(* Logix 5000 project; controller FV vendor 1 type 14 code 217 rev 31.11; software revision 31.00 *)

TASK _1Sec (periodic, rate 1000 ms, priority 10, watchdog 500 ms) : _1Second
TASK MainTask (continuous, watchdog 500 ms) : First_Task, FV_Common, FR_Common, Last_Task

MODULES
   Local : vendor 1 type 14 code 217 (5069 0, rev 31.11)
      MV : vendor 1 type 14 code 217 (Ethernet 192.168.20.32, rev 31.1)
      Remote_IO : vendor 1 type 12 code 298 (Ethernet 192.168.1.1, rev 1.1)
          : vendor 1 type 7 code 82 (Compact 6, rev 1.1, Input RPI 20 ms)
          : vendor 1 type 7 code 76 (Compact 7, rev 1.1, Input RPI 20 ms)
          : vendor 1 type 10 code 47 (Compact 8, rev 1.1, Output RPI 80 ms)
          : 1769-OW16 (Compact 1, rev 1.1, Output RPI 20 ms)
          : 1769-OW16 (Compact 3, rev 1.1, Output RPI 20 ms)
          : 1769-IF8 (Compact 13, rev 1.1, Output RPI 80 ms)
          : 1769-OW16 (Compact 4, rev 1.1, Output RPI 20 ms)
          : 1769-IF8 (Compact 11, rev 1.1, Output RPI 80 ms)
          : 1769-IF8 (Compact 10, rev 1.1, Output RPI 80 ms)
          : 1769-OW16 (Compact 2, rev 1.1, Output RPI 20 ms)
          : 1769-OW16 (Compact 5, rev 1.1, Output RPI 20 ms)
          : 1769-IF8 (Compact 12, rev 1.1, Output RPI 80 ms)
          : vendor 1 type 7 code 79 (Compact 9, rev 3.1, Output RPI 20 ms)
      RIO_Rack_2 : vendor 1 type 12 code 298 (Ethernet 192.168.1.2, rev 1.1)
          : vendor 1 type 7 code 76 (Compact 6, rev 1.1, Input RPI 20 ms)
          : vendor 1 type 7 code 76 (Compact 3, rev 1.1, Input RPI 20 ms)
          : vendor 1 type 7 code 76 (Compact 4, rev 1.1, Input RPI 20 ms)
          : vendor 1 type 7 code 76 (Compact 7, rev 1.1, Input RPI 20 ms)
          : vendor 1 type 7 code 76 (Compact 9, rev 1.1, Input RPI 20 ms)
          : vendor 1 type 7 code 76 (Compact 10, rev 1.1, Input RPI 20 ms)
          : vendor 1 type 7 code 76 (Compact 12, rev 1.1, Input RPI 20 ms)
          : vendor 1 type 7 code 79 (Compact 8, rev 3.1, Output RPI 20 ms)
          : vendor 1 type 10 code 48 (Compact 1, rev 1.1, Output RPI 80 ms)
          : vendor 1 type 10 code 47 (Compact 2, rev 1.1, Output RPI 80 ms)
          : vendor 1 type 7 code 79 (Compact 5, rev 3.1, Output RPI 20 ms)
          : vendor 1 type 7 code 79 (Compact 11, rev 3.1, Output RPI 20 ms)
      RIO_Rack_3 : vendor 1 type 12 code 298 (Ethernet 192.168.1.3, rev 1.1)
          : 1769-IQ16 (Compact 1, rev 1.1, Input RPI 20 ms)
          : 1769-IQ16 (Compact 2, rev 1.1, Input RPI 20 ms)
          : 1769-OW16 (Compact 3, rev 1.1, Output RPI 20 ms)
END_MODULES

TYPE CHECKWORD_FLAGS :   // Checkword Flags
STRUCT
   AUTODRV : DINT;   // Auto-Drive Bit No.
   CLOSEDFB : DINT;   // Closed Feedback Bit No.
   OPENFB : DINT;   // Open Feedback Bit No.
   OUTPUT : DINT;   // Output Bit No.
   MANDRV : DINT;   // Manual Drive Bit No.
   MANUAL : DINT;   // Manual Control Bit No.
   CHECKOFF : DINT;   // Checking Off Bit No.
   TRIPPED : DINT;   // Tripped Bit No.
   FAULT : DINT;   // Fault Bit No.
   SIMFAIL : DINT;   // Simulate Failure Bit
   PREVSCAN : DINT;   // Previous Scan State
   FAULTLOGGED : DINT;   // Fault Logged Flag From Scada
   HIGHLIGHT : DINT;   // Highlight on Graphics
   RUNFB : DINT;   // Pump/Drive Run Feedback
   HEALTHYFB : DINT;   // Pump Healthy Feedback
   NOTTRIPPEDFB : DINT;   // Pump Not Tripped Feedback
   HEALTHYFAULTLOGGED : DINT;   // Pump Not Healthy Fault Logged
   TRIPPEDFAULTLOGGED : DINT;   // Pump Tripped Fault Logged
   INPUTSTATUS : DINT;   // Bit Number for Digital Input Status
   INPUTSTATUSDEBOUNCED : DINT;   // Bit Number For Debounced Input Status
   ANALOGSIMULATION : DINT;   // Bit Number For Analog Simulation Enabled, Used By FactoryTalk
END_STRUCT
END_TYPE

TYPE DateTime :
STRUCT
   Year : DINT;
   Month : DINT;
   Day : DINT;
   Hour : DINT;
   Minute : DINT;
   Second : DINT;
   Microsecond : DINT;
END_STRUCT
END_TYPE

TYPE PlantItem :   // Plant Item
STRUCT
   CW : DINT;   // Checkword
   CheckTime : DINT;   // Check Time
   CheckTimer : DINT;   // Check Time Timer
   DebounceTime : DINT;   // Debounce Time
   DebounceTimer : DINT;   // Debounce Timer
   DriveBits : DINT;   // Item Automatic Drive Bits
   Scaled : REAL;   // Analogue Value Scaled For Input/Output
   RawInput : REAL;   // Raw Input Copied for display On Factory Talk
END_STRUCT
END_TYPE

TYPE Process :   // Data Type For Processes
STRUCT
   Status : DINT;   // Process Current Status
   Step : DINT;   // Process Current Step
   Step_Timer : DINT;   // Current Step Timer
   Fault : DINT;   // Process Current Fault
   Cmd : DINT;   // Command From Scada
   Cmd_avail : DINT;   // Commands Available To Scada
   Cmd_ok : BOOL;   // Startup Command Is Valid Flag
   Cmd_reset : TIMER;   // Startup timer for Invalid Command
   Data_scada : REAL[50];   // Data from Scada
   Data_work : REAL[50];   // Working Data in use by PLC
   Drivebit : DINT;   // Bit Number to Drive Plant Items With
   MessageID : DINT;   // ID to pass with Events/Alarms to Scada
   Past_Prestart : BOOL;   // Flag Set to Indicate past pre start checks.
   Restart_Step : DINT;   // Step to go back to after Continue
END_STRUCT
END_TYPE

TYPE Route :
STRUCT
   CW : DINT;   // Checking Group CW
   CW_Itm : DINT;   // Checking Group Which Has Failed
   Operation : DINT;   // Checking Group Operation Reservation
END_STRUCT
END_TYPE

ADD_ON_INSTRUCTION DayOfWeek   (* revision 1.0 *)
VAR_INPUT
   Year : DINT; {required}
   Month : DINT; {required}
   Day : DINT; {required}
END_VAR
VAR_OUTPUT
   DOW_Output : DINT; {access Read Only, required}
END_VAR
VAR
   DOW_Day : DINT;
   DOW_Year : DINT;
   DOW_Temp00 : REAL;
   DOW_Century : DINT;
   DOW_Month : DINT;
   DOW_Temp01 : REAL;
   DOW_Temp02 : REAL;
   DOW_Temp03 : DINT;
   DOW_Temp04 : DINT;
   DOW_Temp05 : REAL;
   DOW_Temp06 : DINT;
   DOW_Temp07 : REAL;
   DOW_Temp08 : DINT;
   DOW_Temp09 : REAL;
   DOW_Temp10 : REAL;
   DOW_Temp11 : REAL;
   DOW_Temp12 : REAL;
   DOW_Temp13 : REAL;
   DOW_Temp14 : REAL;
   DOW_Temp15 : REAL;
END_VAR

ROUTINE Logic   (* ladder *)
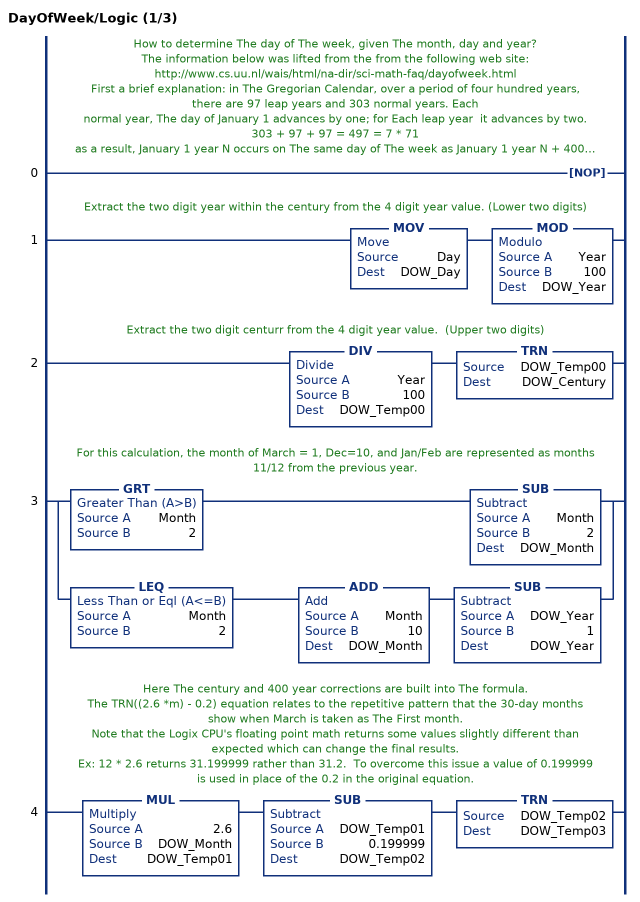
   // How to determine The day of The week, given The month, day and year?
   // The information below was lifted from the from the following web site: http://www.cs.uu.nl/wais/html/na-dir/sci-math-faq/dayofweek.html
   //    First a brief explanation: in The Gregorian Calendar, over a period of four hundred years, there are 97 leap years and 303 normal years. Each
   //  normal year, The day of January 1 advances by one; for Each leap year  it advances by two.
   //    303 + 97 + 97 = 497 = 7 * 71
   //    as a result, January 1 year N occurs on The same day of The week as January 1 year N + 400. Because The leap year pattern also recurs with a four hundred year cycle, a simple table of four hundred elements, and single modulus, suffices to determine The day of The week (in The
   //    Gregorian Calendar), and does it much faster than all The other algorithms proposed. also, Each element takes (in principle) only three bits; The entire table thus takes only 1200 bits; on many computers this will be less than The instructions to do all The complicated calculations proposed or The other algorithms.
   //    Incidental Note: Because 7 does not Divide 400, January 1 occurs more frequently on some days than others! Trick your friends! in a cycle of 400 years, January 1 and March 1 occur on The following days with The following frequencies:
   //            Sun      Mon     Tue     Wed     Thu     Fri     Sat
   //     Jan 1: 58       56      58      57      57      58      56
   //     Mar 1: 58       56      58      56      58      57      57
   //    Of interest is that (contrary to most initial guesses) The occurrence is not maximally flat.
   // In The Mathematical Gazette, vol. 53,, pp.127-129, it is shown that The 13th of The month is more likely to be a Friday than any other day.The author is a 13 year old S.R.Baxter.
   //    The Gregorian Calendar was introduced in 1582 in parts of Europe; it was adopted in 1752 in Great Britain and its colonies, and on various dates in other countries. it replaced The Julian Calendar which has a four-year cycle of leap years; after four years January 1 has advanced by five days. Since 5 is relatively prime to 7, a table of 4 * 7 = 28 elements is necessary for The Julian Calendar.
   //    there is still a 3 day over 10,000 years error which The Gregorian Calendar does not take into account. At some Time such a correction will have to be done but your software will probably not last that long!
   //    Here is a standard method suitable for mental computation:
   //     1. take The last two digits of The year.
   //     2. Divide by 4, discarding any fraction.
   //     3. Add The day of The month.
   //     4. Add The month'S key value: JFM AMJ JAS OND 144 025 036 146
   //     5. Subtract 1 for January or February of a leap year.
   //     6. For a Gregorian Date, Add 0 for 1900'S, 6 for 2000'S, 4 for 1700'S, 2 for 1800'S; for other years, Add or Subtract multiples of 400.
   //     7. For a Julian Date, Add 1 for 1700'S, and 1 for every additional century you go back.
   //     8. Add The last two digits of The year.
   //     9. Divide by 7 and take The remainder.
   //    Now 1 is Sunday, The First day of The week, 2 is Monday, and so on.
   //    The following formula, which is for The Gregorian Calendar only, may be more convenient for computer programming. Note that in some programming languages The remainder operation can yield a negative result if given a negative operand, so mod 7 may not translate to a simple remainder.
   //    W = (k + floor(2.6m - 0.2) - 2C + Y + floor(Y/4) + floor(C/4)) mod 7
   //    where floor() denotes The integer floor function [This is TRN() in Logix],
   // k is day (1 to 31)
   //  m is month (1 = March, ..., 10 = December, 11 = Jan, 12 = Feb) Treat Jan & Feb as months of The preceding year
   //    C is century (1987 has C = 19)
   //    Y is year (1987 has Y = 87 except Y = 86 for Jan & Feb)
   //    W is week day (0 = Sunday, ..., 6 = Saturday)
   //    Here The century and 400 year corrections are built into The formula. The floor(2.6m - 0.2) term relates to The repetitive pattern that The 30-day months show when March is taken as The First month.
   //    The following short C program works for a restricted range, it returns 0 for Monday, 1 for Tuesday, etc.
   // dow(m,d,Y){Y-=m<3;return(Y+Y/4-Y/100+Y/400+"-bed=pen+mad."[m]+d)%7;}
   //    The program appeared was posted by sakamoto@sm.sony.co.jp (Tomohiko sakamoto) on comp.lang.c on March 10th, 1993.
   //    a good mnemonic rule to help on The computation of The day of The week is as follows. in any given year The following days come on The same day of The week: 4/4, 6/6, 8/8, 10/10, 12/12  to remember The next four, remember that I work from 9-5 At a 7-11 so 9/5, 5/9, 7/11, 11/7 and The last day of Feb.
   //    "in 1995 they come on Tuesday. every year this advances one other than leap-years which advance 2. Therefore for 1996 The day will be Thursday, and for 1997 it will be Friday. Therefore ordinarily every 4 years it advances 5 days. there is a minor correction for The century Since The century is a leap year iff The century is divisible by 4. Therefore 2000 is a leap year, but 1900, 1800, and 1700 were not."
   //    Even ignoring The pattern over for a period of years this is still useful Since you can generally figure out what day of The week a given Date is  on faster than someone else can look it up with a calender if The calender is not right there. (a useful skill that.)
   //  References:
   //    Winning Ways for your Mathematical plays. Elwyn R. Berlekamp, John H.  Conway, and Richard k. Guy London ; Toronto : Academic Press, 1982.
   //    Mathematical Carnival. Martin Gardner. New York : Knopf, c1975.
   //    Elementary Number Theory and its applications. Kenneth Rosen. Reading,  Mass. ; Don Mills, Ont. : Addison-Wesley Pub. Co., c1993. p. 156.
   //    Michael Keith and Tom Craver. The Ultimate Perpetual Calendar? Journal of Recreational Mathematics, 22:4, pp. 280-282, 19
   0: NOP();
   // Extract the two digit year within the century from the 4 digit year value. (Lower two digits)
   1: MOV(Day,DOW_Day)MOD(Year,100,DOW_Year);
   // Extract the two digit centurr from the 4 digit year value.  (Upper two digits)
   2: DIV(Year,100,DOW_Temp00)TRN(DOW_Temp00,DOW_Century);
   // For this calculation, the month of March = 1, Dec=10, and Jan/Feb are represented as months 11/12 from the previous year.
   3: [GRT(Month,2) SUB(Month,2,DOW_Month) ,LEQ(Month,2) ADD(Month,10,DOW_Month) SUB(DOW_Year,1,DOW_Year) ];
   // Here The century and 400 year corrections are built into The formula.
   // The TRN((2.6 *m) - 0.2) equation relates to the repetitive pattern that the 30-day months show when March is taken as The First month.
   // Note that the Logix CPU's floating point math returns some values slightly different than expected which can change the final results.
   // Ex: 12 * 2.6 returns 31.199999 rather than 31.2.  To overcome this issue a value of 0.199999 is used in place of the 0.2 in the original equation.
   4: MUL(2.6,DOW_Month,DOW_Temp01)SUB(DOW_Temp01,0.199999,DOW_Temp02)TRN(DOW_Temp02,DOW_Temp03);
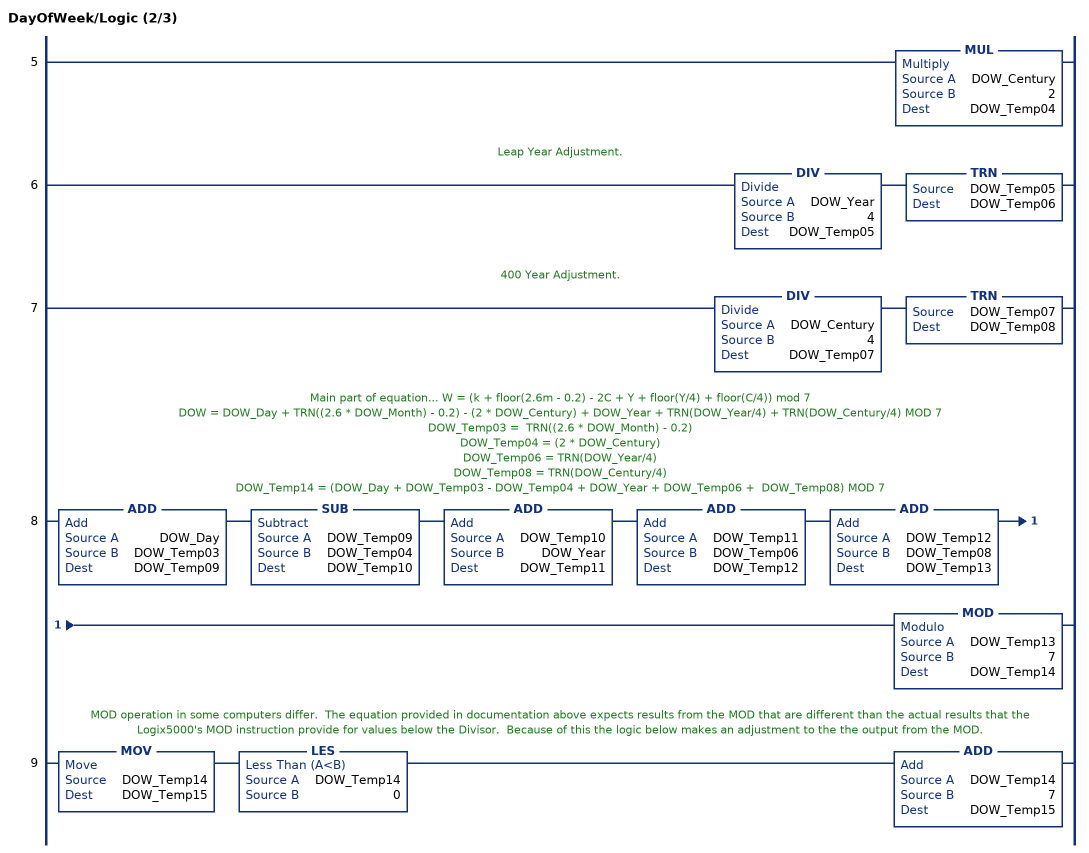
   5: MUL(DOW_Century,2,DOW_Temp04);
   // Leap Year Adjustment.
   6: DIV(DOW_Year,4,DOW_Temp05)TRN(DOW_Temp05,DOW_Temp06);
   // 400 Year Adjustment.
   7: DIV(DOW_Century,4,DOW_Temp07)TRN(DOW_Temp07,DOW_Temp08);
   // Main part of equation... W = (k + floor(2.6m - 0.2) - 2C + Y + floor(Y/4) + floor(C/4)) mod 7
   // DOW = DOW_Day + TRN((2.6 * DOW_Month) - 0.2) - (2 * DOW_Century) + DOW_Year + TRN(DOW_Year/4) + TRN(DOW_Century/4) MOD 7
   // DOW_Temp03 =  TRN((2.6 * DOW_Month) - 0.2)
   // DOW_Temp04 = (2 * DOW_Century)
   // DOW_Temp06 = TRN(DOW_Year/4)
   // DOW_Temp08 = TRN(DOW_Century/4)
   // DOW_Temp14 = (DOW_Day + DOW_Temp03 - DOW_Temp04 + DOW_Year + DOW_Temp06 +  DOW_Temp08) MOD 7
   8: ADD(DOW_Day,DOW_Temp03,DOW_Temp09)SUB(DOW_Temp09,DOW_Temp04,DOW_Temp10)ADD(DOW_Temp10,DOW_Year,DOW_Temp11)ADD(DOW_Temp11,DOW_Temp06,DOW_Temp12)ADD(DOW_Temp12,DOW_Temp08,DOW_Temp13)MOD(DOW_Temp13,7,DOW_Temp14);
   // MOD operation in some computers differ.  The equation provided in documentation above expects results from the MOD that are different than the actual results that the Logix5000's MOD instruction provide for values below the Divisor.  Because of this the logic below makes an adjustment to the the output from the MOD.
   9: MOV(DOW_Temp14,DOW_Temp15)LES(DOW_Temp14,0)ADD(DOW_Temp14,7,DOW_Temp15);
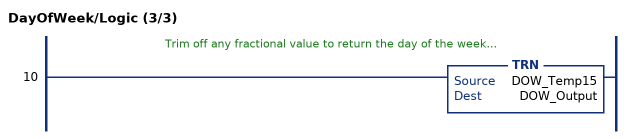
   // Trim off any fractional value to return the day of the week...
   10: TRN(DOW_Temp15,DOW_Output);
END_ROUTINE
END_ADD_ON_INSTRUCTION

VAR_GLOBAL   (* controller tags *)
   _1s_pulse : BOOL;
   Alarm_Reset : BOOL;
   Always_Off : BOOL;
   Always_On : BOOL := 1;
   Analog_Fault_No : DINT := 30001;
   Analog_Simulation_Enabled : BOOL;
   CheckTimeMask : INT := 240;
   CLOCK_system_set : BOOL;
   CLOCKsetvalues : DINT[7] := ([0] := 2019, [1] := 3, [2] := 4, [3] := 6, [5] := 29);
   comms_to_blunger_write_enabled : BOOL;
   comms_to_fv_route_write_enabled : BOOL := 1;
   comms_to_mc_write_enabled : BOOL := 1;
   comms_to_mv_route_write_enabled : BOOL := 1;
   CurrentTime : DateTime := (Year := 2020, Month := 8, Day := 5, Hour := 13, Minute := 9, Second := 51, Microsecond := 283353);
   CWD : CHECKWORD_FLAGS := (CLOSEDFB := 4, OPENFB := 3, OUTPUT := 7, MANDRV := 5, MANUAL := 6, CHECKOFF := 8, FAULT := 15, SIMFAIL := 2, PREVSCAN := 1, FAULTLOGGED := 14, HIGHLIGHT := 9, RUNFB := 3, HEALTHYFB := 10, NOTTRIPPEDFB := 11, HEALTHYFAULTLOGGED := 16, TRIPPEDFAULTLOGGED := 17, INPUTSTATUSDEBOUNCED := 18, ANALOGSIMULATION := 12);
   Default_Check_Time : DINT := 10;
   Delphi_Does_Eng_Func : BOOL;
   Dummy : BOOL := 1;
   FR_0DB : ALIAS FOR FR_B240[0].14;   // 0 0 Debounced
   FR_ALARM_RETURNED_STRING : STRING;
   FR_AUDI1 : PlantItem := (CheckTime := 10);   // AUDI1
   FR_AUDI1_RawOutput : ALIAS FOR RIO_Rack_2:11:O.Data.30;   // FR_AUDI1
   FR_B230 : INT[255] := ([0] := 1);   // FLOW_BITS Flow Meter Bits
        [0].0   // Paraflow flowmeter flow pulse signal One Shot Latch
        [0].1   // Paraflow flowmeter flow pulse signal One Shot Pulse
        [0].2   // Centrifuge1 flowmeter flow pulse signal One Shot Latch
        [0].3   // Centrifuge1 flowmeter flow pulse signal One Shot Pulse
        [0].4   // Centrifuge2 flowmeter flow pulse signal One Shot Latch
        [0].5   // Centrifuge2 flowmeter flow pulse signal One Shot Pulse
   FR_B240 : INT[255] := ([0] := 12944);   // DEBOUNCE Debounce Flags
        [0].0   // FV26/HLP01 FV26 High Level Debounced
        [0].1   // FV26/LLP01 FV26 Low Level Debounced
        [0].10   // FV31/LLP01 FV31 High Level Debounced
        [0].11   // FV31/HLP01 FV31 Low Level Debounced
        [0].12   // VB4/LP01 VB4 Vent level Debounced
        [0].13   // FRV1/LP01 Filtrate Return Vess Level Probe Debounced
        [0].14   // 0 0 Debounced
        [0].15   // 0 0 Debounced
        [0].2   // FV27/HLP01 FV27 High Level Debounced
        [0].3   // FV27/LLP01 FV27 Low Level Debounced
        [0].4   // FV28/HLP01 FV28 High Level Debounced
        [0].5   // FV28/LLP01 FV28 Low Level Debounced
        [0].6   // FV29/HLP01 FV29 High Level Debounced
        [0].7   // FV29/LLP01 FV29 Low Level Debounced
        [0].8   // FV30/LLP01 FV30 High Level Debounced
        [0].9   // FV30/HLP01 FV30 Low Level Debounced
        [1].0   // 0 0 Debounced
        [1].1   // 0 0 Debounced
        [1].10   // 0 0 Debounced
        [1].11   // 0 0 Debounced
        [1].12   // 0 0 Debounced
        [1].13   // 0 0 Debounced
        [1].14   // PanelEstop Panel emergency stop Debounced
        [1].15   // Pilz Pilz healthy input Debounced
        [1].2   // 0 0 Debounced
        [1].3   // 0 0 Debounced
        [1].4   // 0 0 Debounced
        [1].5   // 0 0 Debounced
        [1].6   // 0 0 Debounced
        [1].7   // 0 0 Debounced
        [1].8   // 0 0 Debounced
        [1].9   // 0 0 Debounced
   FR_B246 : INT[255];   // V_REVERSE Flags for reversing contol action
        [0].0   // CLOSE --- VB1/AV08 VB1 Filling Main Block Valve (Reverse Acting)
        [0].1   // CLOSE --- VB2/AV05 VB2 Filling Main Block Valve (Reverse Acting)
        [0].2   // CLOSE FV26/AV01 FV26 Filtrate Inlet Sprayball Bypass CW8
        [0].3   // CLOSE FV27/AV01 FV27 Filtrate Inlet Sprayball Bypass CW13
        [0].4   // CLOSE FV28/AV01 FV28 Filtrate Inlet Sprayball Bypass CW27
        [0].5   // CLOSE FV29/AV01 FV29 Filtrate Inlet Sprayball Bypass CW32
        [0].6   // CLOSE FV30/AV01 FV30 Filtrate Inlet Sprayball Bypass CW64
        [0].7   // CLOSE FV31/AV01 FV31 Filtrate Inlet Sprayball Bypass CW69
        [0].8   // CLOSE --- VB3/AV05 VB3 Filling Main Block Valve (Reverse Acting)
   FR_B247 : INT[255];   // CHECKWORD Simulation Flags for Checkwords
        [0].5   // Checking timebase too short Alarm Increase Timebase OR Number of items to check each timebase
        [0].6   // Do NOT Simulate this item
        [0].7   // Simulate this item
   FR_B248 : INT[255];   // FORCE ON Force On Flags
   FR_B249 : INT[255];   // FORCE_OFF NOT Force Off Flags
   FR_B3 : INT[255] := ([0] := 16, [4] := 1, [7] := 1);   // BINARY
        [0].10   // Disable GEA watchdog
        [0].11   // GEA watchdog fault
        [0].8   // Flowmeter Pulses OSR
        [4].0   // To GEA via MVRoute
        [4].1   // To GEA direct
        [7].0   // YEAST PUMP RUNNING ONE SHOT
   FR_BEACON1 : PlantItem := (CheckTime := 10);   // BEACON1
   FR_BEACON1_RawOutput : ALIAS FOR RIO_Rack_2:11:O.Data.31;   // FR_BEACON1
   FR_bit_data_file_address : DINT;
   FR_bit_file_bit_offset : DINT;
   FR_bit_file_word_offset : DINT;
   FR_bit_offset : DINT;
   FR_bit_returned : BOOL;
   FR_bit_value_to_set : DINT;
   FR_CFG1_P : PlantItem;   // CFG1_P
   FR_CFG1_P_RawInput : ALIAS FOR RIO_Rack_2:12:I.Data.0;   // FR_CFG1_P
   FR_CFG2_P : PlantItem;   // CFG2_P
   FR_CFG2_P_RawInput : ALIAS FOR RIO_Rack_2:12:I.Data.1;   // FR_CFG2_P
   fr_chk_temp : DINT := 2011;
   fr_comms_from_mv_route : MESSAGE;
        MessageParameters(ServiceCode := 16#004c, LocalElement := FR_N13[0], ...)
   fr_comms_from_mv_route2 : MESSAGE;
   fr_comms_from_mvfv_cip : MESSAGE;
        MessageParameters(ServiceCode := 16#004c, LocalElement := FR_N14[0], ...)
   fr_comms_to_MC : MESSAGE;
        MessageParameters(ServiceCode := 16#0faa, LocalElement := FR_N14[100], ...)
   fr_comms_to_MC_timer : TIMER := (PRE := 4000, ACC := 2020, EN := 1, TT := 1);
   fr_comms_to_mv_route : MESSAGE;
        MessageParameters(ServiceCode := 16#0faa, LocalElement := FR_N13[100], ...)
   fr_comms_to_mv_route_timer : TIMER := (PRE := 2000, ACC := 431, EN := 1, TT := 1);
   FR_copy_how_many : DINT;
   FR_Crop_Event_Prefix : STRING := ' FV8 ';
   FR_Crop_Log_ID : DINT := 20;
   FR_data_file_address : DINT := 160;
   FR_data_file_value_to_move : DINT := -1;
   FR_DEFOAM : PlantItem;   // DEFOAM
   FR_DEFOAM_RawOutput : ALIAS FOR RIO_Rack_2:5:O.Data.6;   // FR_DEFOAM
   FR_DEFOAMER : PlantItem;   // DEFOAMER
   FR_DEFOAMER_RawInput : ALIAS FOR RIO_Rack_2:4:I.Data.6;   // FR_DEFOAMER
   FR_Delphi_I : DINT[60] := ([10] := 19823, [11] := 51456, [14] := 1040, [30] := 64);
   FR_Delphi_O : DINT[60] := ([29] := 6144);
   FR_dow_addon_tag : DayOfWeek := (Year := 2020, Month := 8, Day := 5, DOW_Output := 3);
   FR_dow_timer : TIMER := (PRE := 900000, ACC := 788505, EN := 1, TT := 1);
   FR_Event_Alarm_Tag : ALARM_DIGITAL;
   FR_Event_control_FIFO : CONTROL := (LEN := 30, EM := 1);
   FR_Event_control_FIFO_Operation_Type : CONTROL := (LEN := 30, EM := 1);
   FR_Event_Delay_For_Data : TIMER := (PRE := 1000);
   FR_Event_Delay_For_PLC_Startup_Data : TIMER := (PRE := 1000);
   FR_Event_Delay_Timer : TIMER := (PRE := 1000);
   FR_Event_Delay_Timer_Off : TIMER := (PRE := 1000);
   FR_Event_from_buffer : STRING := 'FV 26 Filling Beer Transfer Complete selected by operator (Seb_K)';
   FR_Event_from_buffer_LogData1 : REAL;
   FR_Event_from_buffer_LogData2 : REAL := 226.0;
   FR_Event_from_buffer_LogData3 : REAL;
   FR_Event_from_buffer_LogData4 : REAL;
   FR_Event_from_buffer_Operation_Type : DINT := 22;
   FR_event_step : DINT;
   FR_Event_String_Last : STRING := 'FV 26 Filling Beer Transfer Complete selected by operator (Seb_K)';
   FR_Event_Transact_Trigger_Tag : DINT;
   FR_Events_FIFO_Buffer : STRING[31];
   FR_Events_FIFO_Buffer_Operation_Type : DINT[31];
   FR_F102 : REAL[20] := ([0] := 1.0);
   FR_F202 : REAL[20] := ([0] := 1.032, [1] := 999.0, [2] := 0.28, [3] := 1.0, [4] := 9.81, [5] := 0.8794799, [6] := 0.8794799, [7] := 1.0, [8] := 0.7, [9] := 1.72059);
   FR_F203 : REAL[40] := ([1] := 999.0, [2] := 0.28, [3] := 1.0, [4] := 9.81, [5] := 7.794, [6] := 8.392, [7] := 1.6, [8] := 2.715, [9] := 52.925606, [10] := 3.141, [11] := 9.81, [12] := 0.58931863, [13] := 0.34729645, [14] := 70.42567, [15] := 591.0122, [16] := 7.3712244, [17] := 20.012873, [18] := 67.479744, [19] := 14.554135, [20] := 2.5600002, [21] := 67.479744, [22] := 14.554138, [23] := 51.48848, [24] := 0.6);
   FR_Filling_Event_Prefix : STRING := 'FV 26 ';
   FR_Filling_Log_ID : DINT := 22;
   FR_FILT_PR_PX : PlantItem := (CW := 2#0000_0000_0000_0000_0000_0000_0010_0000);   // FILT_PR_PX
   FR_FILT_PR_PX_RawInput : ALIAS FOR RIO_Rack_2:3:I.Data.25;   // FR_FILT_PR_PX
   FR_FILT_TNK_PX : PlantItem;   // FILT_TNK_PX
   FR_FILT_TNK_PX_RawInput : ALIAS FOR RIO_Rack_2:3:I.Data.26;   // FR_FILT_TNK_PX
   FR_FILT_TNLN_PX : PlantItem := (CW := 2#0000_0000_0000_0100_0000_0000_0000_0001);   // FILT_TNLN_PX
   FR_FILT_TNLN_PX_RawInput : ALIAS FOR RIO_Rack_2:3:I.Data.27;   // FR_FILT_TNLN_PX
   FR_Filtrate_Event_Prefix : STRING := 'FV 27 ';
   FR_Filtrate_Log_ID : DINT := 21;
   FR_from_data_file : DINT := 130;
   FR_from_data_offset : DINT := 110;
   FR_FRV1_AV01 : PlantItem := (CW := 2#0000_0000_0000_0000_0000_0001_1001_0011, CheckTime := 10, CheckTimer := 10, DriveBits := 1);   // FRV1_AV01
   FR_FRV1_AV01_ALARM : ALARM_DIGITAL;
   FR_FRV1_AV01_C : ALIAS FOR RIO_Rack_2:4:I.Data.15;
   FR_FRV1_AV01_DR : ALIAS FOR RIO_Rack_2:5:O.Data.7;
   FR_FRV1_AV01_O : ALIAS FOR RIO_Rack_2:4:I.Data.11;
   FR_FRV1_LP01 : PlantItem := (CW := 2#0000_0000_0000_0000_0000_0000_0010_0000);   // FRV1_LP01
   FR_FRV1_LP01_RawInput : ALIAS FOR RIO_Rack_2:3:I.Data.13;   // FR_FRV1_LP01
   FR_FRV1_LP01DB : ALIAS FOR FR_B240[0].13;   // FRV1/LP01 Filtrate Return Vess Level Probe Debounced
   FR_FV26_AV01 : PlantItem := (CW := 2#0000_0000_0000_0000_0000_0000_0000_1000, CheckTime := 16, CheckTimer := 16);   // FV26_AV01
   FR_FV26_AV01_ALARM : ALARM_DIGITAL;
   FR_FV26_AV01_C : ALIAS FOR RIO_Rack_2:4:I.Data.20;
   FR_FV26_AV01_O : ALIAS FOR RIO_Rack_2:4:I.Data.16;
   FR_FV26_AV01_RDR : ALIAS FOR RIO_Rack_2:5:O.Data.8;
   FR_FV26_AV04 : PlantItem := (CW := 2#0000_0000_0000_0000_0000_0000_0001_0000, CheckTime := 10, CheckTimer := 10);   // FV26_AV04
   FR_FV26_AV04_ALARM : ALARM_DIGITAL;
   FR_FV26_AV04_C : ALIAS FOR RIO_Rack_2:4:I.Data.21;
   FR_FV26_AV04_DR : ALIAS FOR RIO_Rack_2:5:O.Data.9;
   FR_FV26_AV04_O : ALIAS FOR RIO_Rack_2:4:I.Data.17;
   FR_FV26_AV05 : PlantItem := (CW := 2#0000_0000_0000_0000_0000_0000_0001_0000, CheckTime := 10, CheckTimer := 10);   // FV26_AV05
   FR_FV26_AV05_ALARM : ALARM_DIGITAL;
   FR_FV26_AV05_C : ALIAS FOR RIO_Rack_2:4:I.Data.22;
   FR_FV26_AV05_DR : ALIAS FOR RIO_Rack_2:5:O.Data.10;
   FR_FV26_AV05_O : ALIAS FOR RIO_Rack_2:4:I.Data.18;
   FR_FV26_AV06 : PlantItem := (CW := 2#0000_0000_0000_0000_0000_0000_0001_0000, CheckTime := 10, CheckTimer := 10);   // FV26_AV06
   FR_FV26_AV06_ALARM : ALARM_DIGITAL;
   FR_FV26_AV06_C : ALIAS FOR RIO_Rack_2:4:I.Data.23;
   FR_FV26_AV06_DR : ALIAS FOR RIO_Rack_2:5:O.Data.11;
   FR_FV26_AV06_O : ALIAS FOR RIO_Rack_2:4:I.Data.19;
   FR_FV26_AV07 : PlantItem := (CW := 2#0000_0000_0000_0000_0000_0000_0001_0000, CheckTime := 10, CheckTimer := 10);   // FV26_AV07
   FR_FV26_AV07_ALARM : ALARM_DIGITAL;
   FR_FV26_AV07_C : ALIAS FOR RIO_Rack_2:4:I.Data.28;
   FR_FV26_AV07_DR : ALIAS FOR RIO_Rack_2:5:O.Data.12;
   FR_FV26_AV07_O : ALIAS FOR RIO_Rack_2:4:I.Data.24;
   FR_FV26_AV08 : PlantItem := (CW := 2#0000_0000_0000_0000_0000_0000_0001_0000, CheckTime := 16, CheckTimer := 16);   // FV26_AV08
   FR_FV26_AV08_ALARM : ALARM_DIGITAL;
   FR_FV26_AV08_C : ALIAS FOR RIO_Rack_2:12:I.Data.20;
   FR_FV26_AV08_DR : ALIAS FOR FV26_AV08_DUMMY_DR;
   FR_FV26_AV08_O : ALIAS FOR RIO_Rack_2:12:I.Data.16;
   FR_FV26_HLP01 : PlantItem := (CW := 2#0000_0000_0000_0100_0000_0000_0010_0001);   // FV26_HLP01
   FR_FV26_HLP01_RawInput : ALIAS FOR RIO_Rack_2:3:I.Data.0;   // FR_FV26_HLP01
   FR_FV26_HLP01DB : ALIAS FOR FR_B240[0].0;   // FV26/HLP01 FV26 High Level Debounced
   FR_FV26_LLP01 : PlantItem := (CW := 2#0000_0000_0000_0100_0000_0000_0000_0001);   // FV26_LLP01
   FR_FV26_LLP01_RawInput : ALIAS FOR RIO_Rack_2:3:I.Data.1;   // FR_FV26_LLP01
   FR_FV26_LLP01DB : ALIAS FOR FR_B240[0].1;   // FV26/LLP01 FV26 Low Level Debounced
   FR_FV26_LTX01_AI : PlantItem := (CW := 2#0000_0000_0000_0000_1000_0000_0000_0000, CheckTime := 15, CheckTimer := 15, Scaled := 669.40576, RawInput := 7692.0);   // FV26_LTX01
   FR_FV26_LTX01_AI_RawInput : ALIAS FOR RIO_Rack_2:2:I.Ch01Data;   // Real Analog Input , Do Not Use In Code
   FR_FV26_LTX01S : ALIAS FOR FR_N200[10];   // FV26/LTX01 FV26 level transmitter
   FR_FV26_PTX01_AI : PlantItem := (CW := 2#0000_0000_0000_0000_1000_0000_0000_0000, CheckTime := 15, CheckTimer := 15, Scaled := 1.6318126, RawInput := 4009.0);   // FV26_PTX01
   FR_FV26_PTX01_AI_RawInput : ALIAS FOR RIO_Rack_2:2:I.Ch00Data;   // Real Analog Input , Do Not Use In Code
   FR_FV26_PTX01S : ALIAS FOR FR_N200[0];   // FV26/PTX01 FV26 top pressure transmitter
   FR_FV26_ROTO : PlantItem;   // FV26_ROTO
   FR_FV26_ROTO_RawInput : ALIAS FOR RIO_Rack_2:12:I.Data.10;   // FR_FV26_ROTO
   FR_FV26_VA01 : PlantItem := (CheckTime := 10);   // FV26_VA01
   FR_FV26_VA01_RawOutput : ALIAS FOR RIO_Rack_2:11:O.Data.24;   // FR_FV26_VA01
   FR_FV27_AV01 : PlantItem := (CW := 2#0000_0000_0000_0000_0000_0000_0000_1000, CheckTime := 16, CheckTimer := 16);   // FV27_AV01
   FR_FV27_AV01_ALARM : ALARM_DIGITAL;
   FR_FV27_AV01_C : ALIAS FOR RIO_Rack_2:4:I.Data.29;
   FR_FV27_AV01_O : ALIAS FOR RIO_Rack_2:4:I.Data.25;
   FR_FV27_AV01_RDR : ALIAS FOR RIO_Rack_2:5:O.Data.13;
   FR_FV27_AV04 : PlantItem := (CW := 2#0000_0000_0000_0000_0000_0000_0001_0000, CheckTime := 10, CheckTimer := 10);   // FV27_AV04
   FR_FV27_AV04_ALARM : ALARM_DIGITAL;
   FR_FV27_AV04_C : ALIAS FOR RIO_Rack_2:4:I.Data.30;
   FR_FV27_AV04_DR : ALIAS FOR RIO_Rack_2:5:O.Data.14;
   FR_FV27_AV04_O : ALIAS FOR RIO_Rack_2:4:I.Data.26;
   FR_FV27_AV05 : PlantItem := (CW := 2#0000_0000_0000_0000_0000_0000_0001_0000, CheckTime := 10, CheckTimer := 10);   // FV27_AV05
   FR_FV27_AV05_ALARM : ALARM_DIGITAL;
   FR_FV27_AV05_C : ALIAS FOR RIO_Rack_2:4:I.Data.31;
   FR_FV27_AV05_DR : ALIAS FOR RIO_Rack_2:5:O.Data.15;
   FR_FV27_AV05_O : ALIAS FOR RIO_Rack_2:4:I.Data.27;
   FR_FV27_AV06 : PlantItem := (CW := 2#0000_0000_0000_0000_0000_0000_0001_0000, CheckTime := 10, CheckTimer := 10);   // FV27_AV06
   FR_FV27_AV06_ALARM : ALARM_DIGITAL;
   FR_FV27_AV06_C : ALIAS FOR RIO_Rack_2:6:I.Data.4;
   FR_FV27_AV06_DR : ALIAS FOR RIO_Rack_2:5:O.Data.16;
   FR_FV27_AV06_O : ALIAS FOR RIO_Rack_2:6:I.Data.0;
   FR_FV27_AV07 : PlantItem := (CW := 2#0000_0000_0000_0000_0000_0000_0001_0000, CheckTime := 10, CheckTimer := 10);   // FV27_AV07
   FR_FV27_AV07_ALARM : ALARM_DIGITAL;
   FR_FV27_AV07_C : ALIAS FOR RIO_Rack_2:6:I.Data.5;
   FR_FV27_AV07_DR : ALIAS FOR RIO_Rack_2:5:O.Data.17;
   FR_FV27_AV07_O : ALIAS FOR RIO_Rack_2:6:I.Data.1;
   FR_FV27_AV08 : PlantItem := (CW := 2#0000_0000_0000_0000_0000_0000_0001_0000, CheckTime := 16, CheckTimer := 16);   // FV27_AV08
   FR_FV27_AV08_ALARM : ALARM_DIGITAL;
   FR_FV27_AV08_C : ALIAS FOR RIO_Rack_2:12:I.Data.21;
   FR_FV27_AV08_DR : ALIAS FOR FV27_AV08_DUMMY_DR;
   FR_FV27_AV08_O : ALIAS FOR RIO_Rack_2:12:I.Data.17;
   FR_FV27_HLP01 : PlantItem := (CW := 2#0000_0000_0000_0100_0000_0000_0010_0001);   // FV27_HLP01
   FR_FV27_HLP01_RawInput : ALIAS FOR RIO_Rack_2:3:I.Data.2;   // FR_FV27_HLP01
   FR_FV27_HLP01DB : ALIAS FOR FR_B240[0].2;   // FV27/HLP01 FV27 High Level Debounced
   FR_FV27_LLP01 : PlantItem := (CW := 2#0000_0000_0000_0100_0000_0000_0000_0001);   // FV27_LLP01
   FR_FV27_LLP01_RawInput : ALIAS FOR RIO_Rack_2:3:I.Data.3;   // FR_FV27_LLP01
   FR_FV27_LLP01DB : ALIAS FOR FR_B240[0].3;   // FV27/LLP01 FV27 Low Level Debounced
   FR_FV27_LTX01_AI : PlantItem := (CW := 2#0000_0000_0000_0000_1000_0000_0000_0000, CheckTime := 15, CheckTimer := 15, Scaled := 2386.6165, RawInput := 17163.0);   // FV27_LTX01
   FR_FV27_LTX01_AI_RawInput : ALIAS FOR RIO_Rack_2:2:I.Ch03Data;   // Real Analog Input , Do Not Use In Code
   FR_FV27_LTX01S : ALIAS FOR FR_N200[30];   // FV27/LTX01 FV27 level transmitter
   FR_FV27_PTX01_AI : PlantItem := (CW := 2#0000_0000_0000_0000_1000_0000_0000_0000, CheckTime := 15, CheckTimer := 15, Scaled := 1031.1241, RawInput := 9687.0);   // FV27_PTX01
   FR_FV27_PTX01_AI_RawInput : ALIAS FOR RIO_Rack_2:2:I.Ch02Data;   // Real Analog Input , Do Not Use In Code
   FR_FV27_PTX01S : ALIAS FOR FR_N200[20];   // FV27/PTX01 FV27 top pressure transmitter
   FR_FV27_ROTO : PlantItem := (CW := 2#0000_0000_0000_0000_0000_0000_0010_0000);   // FV27_ROTO
   FR_FV27_ROTO_RawInput : ALIAS FOR RIO_Rack_2:12:I.Data.11;   // FR_FV27_ROTO
   FR_FV27_VA01 : PlantItem := (CheckTime := 10);   // FV27_VA01
   FR_FV27_VA01_RawOutput : ALIAS FOR RIO_Rack_2:11:O.Data.25;   // FR_FV27_VA01
   FR_FV28_AV01 : PlantItem := (CW := 2#0000_0000_0000_0000_0000_0000_0000_1000, CheckTime := 16, CheckTimer := 16);   // FV28_AV01
   FR_FV28_AV01_ALARM : ALARM_DIGITAL;
   FR_FV28_AV01_C : ALIAS FOR RIO_Rack_2:6:I.Data.23;
   FR_FV28_AV01_O : ALIAS FOR RIO_Rack_2:6:I.Data.19;
   FR_FV28_AV01_RDR : ALIAS FOR RIO_Rack_2:5:O.Data.27;
   FR_FV28_AV04 : PlantItem := (CW := 2#0000_0000_0000_0000_0000_0000_0001_0000, CheckTime := 10, CheckTimer := 10);   // FV28_AV04
   FR_FV28_AV04_ALARM : ALARM_DIGITAL;
   FR_FV28_AV04_C : ALIAS FOR RIO_Rack_2:6:I.Data.28;
   FR_FV28_AV04_DR : ALIAS FOR RIO_Rack_2:5:O.Data.28;
   FR_FV28_AV04_O : ALIAS FOR RIO_Rack_2:6:I.Data.24;
   FR_FV28_AV05 : PlantItem := (CW := 2#0000_0000_0000_0000_0000_0000_0001_0000, CheckTime := 10, CheckTimer := 10);   // FV28_AV05
   FR_FV28_AV05_ALARM : ALARM_DIGITAL;
   FR_FV28_AV05_C : ALIAS FOR RIO_Rack_2:6:I.Data.29;
   FR_FV28_AV05_DR : ALIAS FOR RIO_Rack_2:5:O.Data.29;
   FR_FV28_AV05_O : ALIAS FOR RIO_Rack_2:6:I.Data.25;
   FR_FV28_AV06 : PlantItem := (CW := 2#0000_0000_0000_0000_0000_0000_0001_0000, CheckTime := 10, CheckTimer := 10);   // FV28_AV06
   FR_FV28_AV06_ALARM : ALARM_DIGITAL;
   FR_FV28_AV06_C : ALIAS FOR RIO_Rack_2:6:I.Data.30;
   FR_FV28_AV06_DR : ALIAS FOR RIO_Rack_2:5:O.Data.30;
   FR_FV28_AV06_O : ALIAS FOR RIO_Rack_2:6:I.Data.26;
   FR_FV28_AV07 : PlantItem := (CW := 2#0000_0000_0000_0000_0000_0000_0011_0000, CheckTime := 10, CheckTimer := 10);   // FV28_AV07
   FR_FV28_AV07_ALARM : ALARM_DIGITAL;
   FR_FV28_AV07_C : ALIAS FOR RIO_Rack_2:6:I.Data.31;
   FR_FV28_AV07_DR : ALIAS FOR RIO_Rack_2:5:O.Data.31;
   FR_FV28_AV07_O : ALIAS FOR RIO_Rack_2:6:I.Data.27;
   FR_FV28_AV08 : PlantItem := (CW := 2#0000_0000_0000_0000_0000_0000_0001_0000, CheckTime := 16, CheckTimer := 16);   // FV28_AV08
   FR_FV28_AV08_ALARM : ALARM_DIGITAL;
   FR_FV28_AV08_C : ALIAS FOR RIO_Rack_2:12:I.Data.22;
   FR_FV28_AV08_DR : ALIAS FOR FV28_AV08_DUMMY_DR;
   FR_FV28_AV08_O : ALIAS FOR RIO_Rack_2:12:I.Data.18;
   FR_FV28_HLP01 : PlantItem := (CW := 2#0000_0000_0000_0000_0000_0000_0010_0000);   // FV28_HLP01
   FR_FV28_HLP01_RawInput : ALIAS FOR RIO_Rack_2:3:I.Data.4;   // FR_FV28_HLP01
   FR_FV28_HLP01DB : ALIAS FOR FR_B240[0].4;   // FV28/HLP01 FV28 High Level Debounced
   FR_FV28_LLP01 : PlantItem := (CW := 2#0000_0000_0000_0100_0000_0000_0000_0001);   // FV28_LLP01
   FR_FV28_LLP01_RawInput : ALIAS FOR RIO_Rack_2:3:I.Data.5;   // FR_FV28_LLP01
   FR_FV28_LLP01DB : ALIAS FOR FR_B240[0].5;   // FV28/LLP01 FV28 Low Level Debounced
   FR_FV28_LTX01_AI : PlantItem := (CW := 2#0000_0000_0000_0000_1000_0000_0000_0000, CheckTime := 15, CheckTimer := 15, Scaled := 1150.2465, RawInput := 10344.0);   // FV28_LTX01
   FR_FV28_LTX01_AI_RawInput : ALIAS FOR RIO_Rack_2:2:I.Ch05Data;   // Real Analog Input , Do Not Use In Code
   FR_FV28_LTX01S : ALIAS FOR FR_N200[50];   // FV28/LTX01 FV28 level transmitter
   FR_FV28_PTX01_AI : PlantItem := (CW := 2#0000_0000_0000_0000_1000_0000_0000_0000, CheckTime := 15, CheckTimer := 15, Scaled := 1.087875, RawInput := 4006.0);   // FV28_PTX01
   FR_FV28_PTX01_AI_RawInput : ALIAS FOR RIO_Rack_2:2:I.Ch04Data;   // Real Analog Input , Do Not Use In Code
   FR_FV28_PTX01S : ALIAS FOR FR_N200[40];   // FV28/PTX01 FV28 top pressure transmitter
   FR_FV28_ROTO : PlantItem := (CW := 2#0000_0000_0000_0000_0000_0000_0010_0000);   // FV28_ROTO
   FR_FV28_ROTO_RawInput : ALIAS FOR RIO_Rack_2:12:I.Data.12;   // FR_FV28_ROTO
   FR_FV28_V : PlantItem := (CheckTime := 10);   // FV28_V
   FR_FV28_V_RawOutput : ALIAS FOR RIO_Rack_2:11:O.Data.20;   // FR_FV28_V
   FR_FV28_VA01 : PlantItem := (CheckTime := 10);   // FV28_VA01
   FR_FV28_VA01_RawOutput : ALIAS FOR RIO_Rack_2:11:O.Data.26;   // FR_FV28_VA01
   FR_FV29_AV01 : PlantItem := (CW := 2#0000_0000_0000_0000_0000_0000_0000_1000, CheckTime := 16, CheckTimer := 16);   // FV29_AV01
   FR_FV29_AV01_ALARM : ALARM_DIGITAL;
   FR_FV29_AV01_C : ALIAS FOR RIO_Rack_2:7:I.Data.4;
   FR_FV29_AV01_O : ALIAS FOR RIO_Rack_2:7:I.Data.0;
   FR_FV29_AV01_RDR : ALIAS FOR RIO_Rack_2:8:O.Data.0;
   FR_FV29_AV04 : PlantItem := (CW := 2#0000_0000_0000_0000_0000_0000_0001_0000, CheckTime := 10, CheckTimer := 10);   // FV29_AV04
   FR_FV29_AV04_ALARM : ALARM_DIGITAL;
   FR_FV29_AV04_C : ALIAS FOR RIO_Rack_2:7:I.Data.5;
   FR_FV29_AV04_DR : ALIAS FOR RIO_Rack_2:8:O.Data.1;
   FR_FV29_AV04_O : ALIAS FOR RIO_Rack_2:7:I.Data.1;
   FR_FV29_AV05 : PlantItem := (CW := 2#0000_0000_0000_0000_0000_0000_0001_0000, CheckTime := 10, CheckTimer := 10);   // FV29_AV05
   FR_FV29_AV05_ALARM : ALARM_DIGITAL;
   FR_FV29_AV05_C : ALIAS FOR RIO_Rack_2:7:I.Data.6;
   FR_FV29_AV05_DR : ALIAS FOR RIO_Rack_2:8:O.Data.2;
   FR_FV29_AV05_O : ALIAS FOR RIO_Rack_2:7:I.Data.2;
   FR_FV29_AV06 : PlantItem := (CW := 2#0000_0000_0000_0000_0000_0000_0001_0000, CheckTime := 10, CheckTimer := 10);   // FV29_AV06
   FR_FV29_AV06_ALARM : ALARM_DIGITAL;
   FR_FV29_AV06_C : ALIAS FOR RIO_Rack_2:7:I.Data.7;
   FR_FV29_AV06_DR : ALIAS FOR RIO_Rack_2:8:O.Data.3;
   FR_FV29_AV06_O : ALIAS FOR RIO_Rack_2:7:I.Data.3;
   FR_FV29_AV07 : PlantItem := (CW := 2#0000_0000_0000_0000_0000_0000_0001_0000, CheckTime := 10, CheckTimer := 10);   // FV29_AV07
   FR_FV29_AV07_ALARM : ALARM_DIGITAL;
   FR_FV29_AV07_C : ALIAS FOR RIO_Rack_2:7:I.Data.12;
   FR_FV29_AV07_DR : ALIAS FOR RIO_Rack_2:8:O.Data.4;
   FR_FV29_AV07_O : ALIAS FOR RIO_Rack_2:7:I.Data.8;
   FR_FV29_AV08 : PlantItem := (CW := 2#0000_0000_0000_0000_0000_0000_0001_0000, CheckTime := 16, CheckTimer := 16);   // FV29_AV08
   FR_FV29_AV08_ALARM : ALARM_DIGITAL;
   FR_FV29_AV08_C : ALIAS FOR RIO_Rack_2:12:I.Data.23;
   FR_FV29_AV08_DR : ALIAS FOR FV29_AV08_DUMMY_DR;
   FR_FV29_AV08_O : ALIAS FOR RIO_Rack_2:12:I.Data.19;
   FR_FV29_HLP01 : PlantItem := (CW := 2#0000_0000_0000_0100_0000_0000_0010_0001);   // FV29_HLP01
   FR_FV29_HLP01_RawInput : ALIAS FOR RIO_Rack_2:3:I.Data.6;   // FR_FV29_HLP01
   FR_FV29_HLP01DB : ALIAS FOR FR_B240[0].6;   // FV29/HLP01 FV29 High Level Debounced
   FR_FV29_LLP01 : PlantItem;   // FV29_LLP01
   FR_FV29_LLP01_RawInput : ALIAS FOR RIO_Rack_2:3:I.Data.7;   // FR_FV29_LLP01
   FR_FV29_LLP01DB : ALIAS FOR FR_B240[0].7;   // FV29/LLP01 FV29 Low Level Debounced
   FR_FV29_LTX01_AI : PlantItem := (CW := 2#0000_0000_0000_0000_1000_0000_0000_0000, CheckTime := 15, CheckTimer := 15, Scaled := -0.72525, RawInput := 3996.0);   // FV29_LTX01
   FR_FV29_LTX01_AI_RawInput : ALIAS FOR RIO_Rack_2:2:I.Ch07Data;   // Real Analog Input , Do Not Use In Code
   FR_FV29_LTX01S : ALIAS FOR FR_N200[70];   // FV29/LTX01 FV29 level transmitter
   FR_FV29_PTX01_AI : PlantItem := (CW := 2#0000_0000_0000_0000_1000_0000_0000_0000, CheckTime := 15, CheckTimer := 15, Scaled := 5.9833126, RawInput := 4033.0);   // FV29_PTX01
   FR_FV29_PTX01_AI_RawInput : ALIAS FOR RIO_Rack_2:2:I.Ch06Data;   // Real Analog Input , Do Not Use In Code
   FR_FV29_PTX01S : ALIAS FOR FR_N200[60];   // FV29/PTX01 FV29 top pressure transmitter
   FR_FV29_ROTO : PlantItem := (CW := 2#0000_0000_0000_0000_0000_0000_0010_0000);   // FV29_ROTO
   FR_FV29_ROTO_RawInput : ALIAS FOR RIO_Rack_2:12:I.Data.13;   // FR_FV29_ROTO
   FR_FV29_VA01 : PlantItem := (CW := 2#0000_0000_0000_0000_0000_0000_1000_0001, CheckTime := 10, DriveBits := 1);   // FV29_VA01
   FR_FV29_VA01_RawOutput : ALIAS FOR RIO_Rack_2:11:O.Data.27;   // FR_FV29_VA01
   FR_FV30_AV01 : PlantItem := (CW := 2#0000_0000_0000_0000_0000_0000_0000_1000, CheckTime := 16, CheckTimer := 16);   // FV30_AV01
   FR_FV30_AV01_ALARM : ALARM_DIGITAL;
   FR_FV30_AV01_C : ALIAS FOR RIO_Rack_2:10:I.Data.4;
   FR_FV30_AV01_O : ALIAS FOR RIO_Rack_2:10:I.Data.0;
   FR_FV30_AV01_RDR : ALIAS FOR RIO_Rack_2:11:O.Data.0;
   FR_FV30_AV04 : PlantItem := (CW := 2#0000_0000_0000_0000_0000_0000_0001_0000, CheckTime := 10, CheckTimer := 10);   // FV30_AV04
   FR_FV30_AV04_ALARM : ALARM_DIGITAL;
   FR_FV30_AV04_C : ALIAS FOR RIO_Rack_2:10:I.Data.5;
   FR_FV30_AV04_DR : ALIAS FOR RIO_Rack_2:11:O.Data.1;
   FR_FV30_AV04_O : ALIAS FOR RIO_Rack_2:10:I.Data.1;
   FR_FV30_AV05 : PlantItem := (CW := 2#0000_0000_0000_0000_0000_0000_0001_0000, CheckTime := 10, CheckTimer := 10);   // FV30_AV05
   FR_FV30_AV05_ALARM : ALARM_DIGITAL;
   FR_FV30_AV05_C : ALIAS FOR RIO_Rack_2:10:I.Data.6;
   FR_FV30_AV05_DR : ALIAS FOR RIO_Rack_2:11:O.Data.2;
   FR_FV30_AV05_O : ALIAS FOR RIO_Rack_2:10:I.Data.2;
   FR_FV30_AV06 : PlantItem := (CW := 2#0000_0000_0000_0000_0000_0000_0001_0000, CheckTime := 10, CheckTimer := 10);   // FV30_AV06
   FR_FV30_AV06_ALARM : ALARM_DIGITAL;
   FR_FV30_AV06_C : ALIAS FOR RIO_Rack_2:10:I.Data.7;
   FR_FV30_AV06_DR : ALIAS FOR RIO_Rack_2:11:O.Data.3;
   FR_FV30_AV06_O : ALIAS FOR RIO_Rack_2:10:I.Data.3;
   FR_FV30_AV07 : PlantItem := (CW := 2#0000_0000_0000_0000_0000_0000_0001_0000, CheckTime := 10, CheckTimer := 10);   // FV30_AV07
   FR_FV30_AV07_ALARM : ALARM_DIGITAL;
   FR_FV30_AV07_C : ALIAS FOR RIO_Rack_2:10:I.Data.12;
   FR_FV30_AV07_DR : ALIAS FOR RIO_Rack_2:11:O.Data.4;
   FR_FV30_AV07_O : ALIAS FOR RIO_Rack_2:10:I.Data.8;
   FR_FV30_AV08 : PlantItem := (CW := 2#0000_0000_0000_0000_0000_0000_0001_0000, CheckTime := 16, CheckTimer := 16);   // FV30_AV08
   FR_FV30_AV08_ALARM : ALARM_DIGITAL;
   FR_FV30_AV08_C : ALIAS FOR RIO_Rack_2:12:I.Data.28;
   FR_FV30_AV08_DR : ALIAS FOR FV30_AV08_DUMMY_DR;
   FR_FV30_AV08_O : ALIAS FOR RIO_Rack_2:12:I.Data.24;
   FR_FV30_HLP01 : PlantItem := (CW := 2#0000_0000_0000_0100_0000_0000_0010_0001);   // FV30_HLP01
   FR_FV30_HLP01_RawInput : ALIAS FOR RIO_Rack_2:3:I.Data.8;   // FR_FV30_HLP01
   FR_FV30_HLP01DB : ALIAS FOR FR_B240[0].9;   // FV30/HLP01 FV30 Low Level Debounced
   FR_FV30_LLP01 : PlantItem := (CW := 2#0000_0000_0000_0000_0000_0000_0010_0000);   // FV30_LLP01
   FR_FV30_LLP01_RawInput : ALIAS FOR RIO_Rack_2:3:I.Data.9;   // FR_FV30_LLP01
   FR_FV30_LLP01DB : ALIAS FOR FR_B240[0].8;   // FV30/LLP01 FV30 High Level Debounced
   FR_FV30_LTX01_AI : PlantItem := (CW := 2#0000_0000_0000_0000_1000_0000_0000_0000, CheckTime := 15, CheckTimer := 15, Scaled := -7.112813, RawInput := 3973.0);   // FV30_LTX01
   FR_FV30_LTX01_AI_RawInput : ALIAS FOR RIO_Rack_2:2:I.Ch09Data;   // Real Analog Input , Do Not Use In Code
   FR_FV30_LTX01S : ALIAS FOR FR_N200[90];   // FV30/LTX01 FV30 level transmitter
   FR_FV30_PTX01_AI : PlantItem := (CW := 2#0000_0000_0000_0000_1000_0000_0000_0000, CheckTime := 15, CheckTimer := 15, Scaled := -4.741875, RawInput := 3982.0);   // FV30_PTX01
   FR_FV30_PTX01_AI_RawInput : ALIAS FOR RIO_Rack_2:2:I.Ch08Data;   // Real Analog Input , Do Not Use In Code
   FR_FV30_PTX01S : ALIAS FOR FR_N200[80];   // FV30/PTX01 FV30 top pressure transmitter
   FR_FV30_ROTO : PlantItem := (CW := 2#0000_0000_0000_0000_0000_0000_0010_0000);   // FV30_ROTO
   FR_FV30_ROTO_RawInput : ALIAS FOR RIO_Rack_2:12:I.Data.14;   // FR_FV30_ROTO
   FR_FV30_VA01 : PlantItem := (CW := 2#0000_0000_0000_0000_0000_0000_1000_0001, CheckTime := 10, DriveBits := 1);   // FV30_VA01
   FR_FV30_VA01_RawOutput : ALIAS FOR RIO_Rack_2:11:O.Data.28;   // FR_FV30_VA01
   FR_FV31_AV01 : PlantItem := (CW := 2#0000_0000_0000_0000_0000_0000_0000_1000, CheckTime := 16, CheckTimer := 16);   // FV31_AV01
   FR_FV31_AV01_ALARM : ALARM_DIGITAL;
   FR_FV31_AV01_C : ALIAS FOR RIO_Rack_2:10:I.Data.13;
   FR_FV31_AV01_O : ALIAS FOR RIO_Rack_2:10:I.Data.9;
   FR_FV31_AV01_RDR : ALIAS FOR RIO_Rack_2:11:O.Data.5;
   FR_FV31_AV04 : PlantItem := (CW := 2#0000_0000_0000_0000_0000_0000_0001_0000, CheckTime := 10, CheckTimer := 10);   // FV31_AV04
   FR_FV31_AV04_ALARM : ALARM_DIGITAL;
   FR_FV31_AV04_C : ALIAS FOR RIO_Rack_2:10:I.Data.14;
   FR_FV31_AV04_DR : ALIAS FOR RIO_Rack_2:11:O.Data.6;
   FR_FV31_AV04_O : ALIAS FOR RIO_Rack_2:10:I.Data.10;
   FR_FV31_AV05 : PlantItem := (CW := 2#0000_0000_0000_0000_0000_0000_0001_0000, CheckTime := 10, CheckTimer := 10);   // FV31_AV05
   FR_FV31_AV05_ALARM : ALARM_DIGITAL;
   FR_FV31_AV05_C : ALIAS FOR RIO_Rack_2:10:I.Data.15;
   FR_FV31_AV05_DR : ALIAS FOR RIO_Rack_2:11:O.Data.7;
   FR_FV31_AV05_O : ALIAS FOR RIO_Rack_2:10:I.Data.11;
   FR_FV31_AV06 : PlantItem := (CW := 2#0000_0000_0000_0000_0000_0000_0001_0000, CheckTime := 10, CheckTimer := 10);   // FV31_AV06
   FR_FV31_AV06_ALARM : ALARM_DIGITAL;
   FR_FV31_AV06_C : ALIAS FOR RIO_Rack_2:10:I.Data.20;
   FR_FV31_AV06_DR : ALIAS FOR RIO_Rack_2:11:O.Data.8;
   FR_FV31_AV06_O : ALIAS FOR RIO_Rack_2:10:I.Data.16;
   FR_FV31_AV07 : PlantItem := (CW := 2#0000_0000_0000_0000_0000_0000_0001_0000, CheckTime := 10, CheckTimer := 10);   // FV31_AV07
   FR_FV31_AV07_ALARM : ALARM_DIGITAL;
   FR_FV31_AV07_C : ALIAS FOR RIO_Rack_2:10:I.Data.21;
   FR_FV31_AV07_DR : ALIAS FOR RIO_Rack_2:11:O.Data.9;
   FR_FV31_AV07_O : ALIAS FOR RIO_Rack_2:10:I.Data.17;
   FR_FV31_AV08 : PlantItem := (CW := 2#0000_0000_0000_0000_0000_0000_0001_0000, CheckTime := 16, CheckTimer := 16);   // FV31_AV08
   FR_FV31_AV08_ALARM : ALARM_DIGITAL;
   FR_FV31_AV08_C : ALIAS FOR RIO_Rack_2:12:I.Data.29;
   FR_FV31_AV08_DR : ALIAS FOR FV31_AV08_DUMMY_DR;
   FR_FV31_AV08_O : ALIAS FOR RIO_Rack_2:12:I.Data.25;
   FR_FV31_HLP01 : PlantItem := (CW := 2#0000_0000_0000_0100_0000_0000_0010_0001);   // FV31_HLP01
   FR_FV31_HLP01_RawInput : ALIAS FOR RIO_Rack_2:3:I.Data.10;   // FR_FV31_HLP01
   FR_FV31_HLP01DB : ALIAS FOR FR_B240[0].11;   // FV31/HLP01 FV31 Low Level Debounced
   FR_FV31_LLP01 : PlantItem := (CW := 2#0000_0000_0000_0100_0000_0000_0000_0001);   // FV31_LLP01
   FR_FV31_LLP01_RawInput : ALIAS FOR RIO_Rack_2:3:I.Data.11;   // FR_FV31_LLP01
   FR_FV31_LLP01DB : ALIAS FOR FR_B240[0].10;   // FV31/LLP01 FV31 High Level Debounced
   FR_FV31_LTX01_AI : PlantItem := (CW := 2#0000_0000_0000_0000_1000_0000_0000_0000, CheckTime := 15, CheckTimer := 15, Scaled := 1142.265, RawInput := 8336.0);   // FV31_LTX01
   FR_FV31_LTX01_AI_RawInput : ALIAS FOR RIO_Rack_2:2:I.Ch11Data;   // Real Analog Input , Do Not Use In Code
   FR_FV31_LTX01S : ALIAS FOR FR_N200[110];   // FV31/LTX01 FV31 level transmitter
   FR_FV31_PTX01_AI : PlantItem := (CW := 2#0000_0000_0000_0000_1000_0000_0000_0000, CheckTime := 15, CheckTimer := 15, Scaled := -1.05375, RawInput := 3996.0);   // FV31_PTX01
   FR_FV31_PTX01_AI_RawInput : ALIAS FOR RIO_Rack_2:2:I.Ch10Data;   // Real Analog Input , Do Not Use In Code
   FR_FV31_PTX01S : ALIAS FOR FR_N200[100];   // FV31/PTX01 FV31 top pressure transmitter
   FR_FV31_ROTO : PlantItem := (CW := 2#0000_0000_0000_0000_0000_0000_0010_0000);   // FV31_ROTO
   FR_FV31_ROTO_RawInput : ALIAS FOR RIO_Rack_2:12:I.Data.15;   // FR_FV31_ROTO
   FR_FV31_VA01 : PlantItem := (CheckTime := 10);   // FV31_VA01
   FR_FV31_VA01_RawOutput : ALIAS FOR RIO_Rack_2:11:O.Data.29;   // FR_FV31_VA01
   FR_FVR1_P01 : PlantItem := (CW := 2#0000_0000_0000_0000_0000_1100_0000_0000, CheckTime := 10, CheckTimer := 15);   // FVR1_P01
   FR_FVR1_P01_ALARM : ALARM_DIGITAL;
   FR_FVR1_P01_D : ALIAS FOR RIO_Rack_2:5:O.Data.5;
   FR_FVR1_P01_R : ALIAS FOR RIO_Rack_2:4:I.Data.9;
   FR_FVs26_31_Cropping_Event : STRING;
   FR_FVs26_31_Filling_Event : STRING;
   FR_FVs26_31_Filtrate_Event : STRING;
   FR_FVs26_31_Green_Beer_Event : STRING;
   FR_FVS_P01 : PlantItem := (CW := 2#0000_0000_0000_0000_0000_1100_0000_0000, CheckTime := 10, CheckTimer := 10);   // FVS_P01
   FR_FVS_P01_ALARM : ALARM_DIGITAL;
   FR_FVS_P01_D : ALIAS FOR RIO_Rack_2:5:O.Data.0;
   FR_FVS_P01_R : ALIAS FOR RIO_Rack_2:4:I.Data.0;
   FR_GBM_P01 : PlantItem := (CW := 2#0000_0000_0000_0000_0000_1100_0000_0000, CheckTime := 10, CheckTimer := 10);   // GBM_P01
   FR_GBM_P01_ALARM : ALARM_DIGITAL;
   FR_GBM_P01_D : ALIAS FOR RIO_Rack_2:5:O.Data.2;
   FR_GBM_P01_R : ALIAS FOR RIO_Rack_2:4:I.Data.2;
   FR_GreenBeer_Event_Prefix : STRING := 'FV 26 ';
   FR_GreenBeer_Log_ID : DINT := 23;
   FR_Last_LogData_For_Op : REAL[30,20] := ([3,2] := 96.0, [4,2] := 26.0, [5,1] := 2.0, [5,2] := 25.0, [6,1] := 28.0, [8,1] := 28.0, [10,1] := 96.0, [20,1] := 8.0, [21,1] := 229.0, [22,2] := 226.0, [23,1] := 226.0);